// TIA Portal project "Demontagestation" (V17) (continued)
VERSION : 0.1
   VAR_INPUT
      Freigeben : Bool;   // "true", wenn der Funktionbaustein ausgeführt werden soll; bei "false werden die Ausgänge auf "Null" gesetzt
      Befehlsindex : USInt;   // Der Index zeigt auf einem Befehl, den der Greifer dann ausführen soll. {0 = FastStop, 1 = Stop, 2 = Quittierung, 3 = Referenzierung, 4 = Hubmessung, 5 = Greifen, 6 = Loslassen, 7 = Positionsfahrt, 8 = Relativfahrt}
      Kraftmodus : USInt;   // Der Wert (0 - 7) stellt die Art (Fast- oder Softgrip) und Kraft (100%, 75%, 50%, 25%) des Greifens ein (relevant bei Greifen).
      Außen_Innen : Bool;   // "true", wenn das Werkstück von innen gegriffen werden soll, sonst "false" (relevant bei Greifen und Loslassen)
      Zielposition : Real;   // Der Geifer positioniert sich nach dem vorgegebenen Positionswert (relevant bei Positions- und Relativfahrt).
   END_VAR
   VAR_OUTPUT
      Rückmeldung : String;   // Detaillierte Informationen über den Ausführungsstatus
      Fehler : Bool;   // "true", wenn im Prozess einen Fehler anliegt
      Fehlermeldung : String;   // Detaillierte Informationen über den Fehler.
      Hub_aktuell : Real;   // Der aktuelle Wert der Postition des Greifers
   END_VAR
   VAR_IN_OUT
      Ausführen : Bool;   // "true", um zu bestätigen, dass der Greifer aus den eingetragenen Daten den Befehl ausführen soll
   END_VAR
   VAR
      Befehlswert : Byte;   // Rohdatenwert eines Befehls
   END_VAR
   VAR_TEMP
      Prozessbit : Bool;   // "true", wenn der Befehl abgearbeitet ist
      Erfolg : Bool;   // "true", wenn der Befehl erfolgreich vollständig ausgeführt wurde
      Error : Bool;   // Quittierungspflichtige Fehler
      Spezifikationsfehler : Bool;   // Fehler, bei dem ein eingetragener Wert außerhalb des Gültigkeitsbereiches liegt
      Wartung : Bool;   // "true", wenn der Greifer gewartet werden muss
      Betrieb : Bool;   // "true", wenn der Greifer betriebsbereit ist
      Referenziert : Bool;   // "true", wenn der Greifer referenziert ist
   END_VAR
   VAR CONSTANT
      "BEGINN_E-ADRESSE" : Int := 39;   // Beginn der Eingangsadresse in Hardware-Konfiguration
      "BEGINN_A-ADRESSE" : Int := 29;   // Beginn der Eingangsadresse in Hardware-Konfiguration / Beginn der Ausgangsadresse in Hardware-Konfiguration
      NOTINDEX : USInt := 0;   // Index, der auf einem Notbefehl zuweist
      FEHLERWERT : Byte := -1;   // Wert, der statt auf einem Befehl einem Fehler weist.
      QUITTIERUNG : Byte := 16#1;   // Nach Beheben eines Fehlers wird der Greifer durch Quittieren des Fehlers vom Fehlerzustand in den normalen Betriebszustand versetzt.
      REFERENZIERUNG : Byte := 16#2;   // Beim Referenzieren wird die Nullposition festgelegt. Der Greifer fährt in eingestellter Referenzierrichtung bis zum mechanischen Endanschlag.
      HUBMESSUNG : Byte := 16#7;   // Bei der Hubmessung wird der maximale Hub des Greifers gegenüber der Referenzierposition festgelegt.
      GREIFEN : Byte := 16#4;   // Beim Greifen wird in Greifrichtung bis zum Anschlag gefahren und das Werkstück mit eingestellter Greifkraft gehalten.
      LOSLASSEN : Byte := 16#3;   // Beim Loslassen wird entgegen der Greifrichtung bis auf Endanschlag gefahren.
      POSITIONSFAHRT : Byte := 16#5;   // Der Geifer fährt auf die unter "Zielposition" angegebene Position.
      RELATIVFAHRT : Byte := 16#6;   // Der Geifer fährt auf eine Position, die von der letzten aktuellen Position mit einem relativen Abstand ermittelt wird.
      STOP : Byte := 16#8;   // Der Greifer wird geregelt in Stillstand versetzt.
      FASTSTOP : Byte := 16#0;   // Die elektrische Energieversorgung zum Aktor wird sofort unterbrochen, der Greifer wird ungesteuert stillgesetzt.
   END_VAR
BEGIN

REGION Network 1: Befehlszuweisung
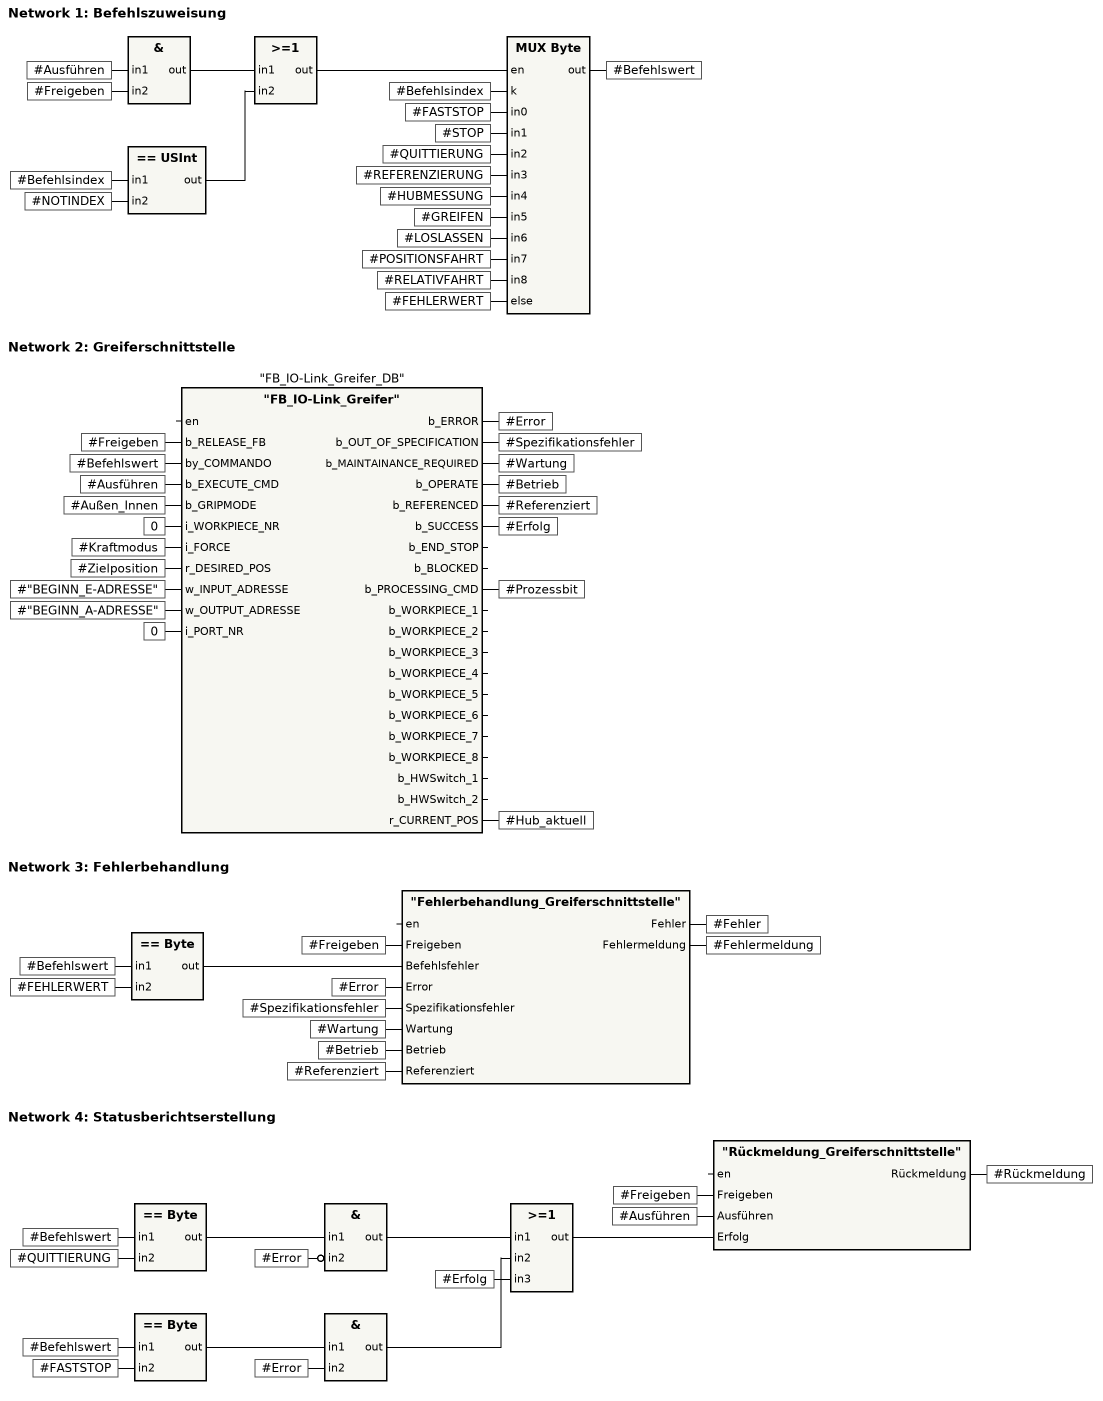
   // no SCL statement known for Mux: written as a call
   IF (#Ausführen AND #Freigeben) OR (#Befehlsindex = #NOTINDEX) THEN
       Mux(k := #Befehlsindex,
           in0 := #FASTSTOP,
           in1 := #STOP,
           in2 := #QUITTIERUNG,
           in3 := #REFERENZIERUNG,
           in4 := #HUBMESSUNG,
           in5 := #GREIFEN,
           in6 := #LOSLASSEN,
           in7 := #POSITIONSFAHRT,
           in8 := #RELATIVFAHRT,
           "else" := #FEHLERWERT,
           out => #Befehlswert);
   END_IF;
END_REGION

REGION Network 2: Greiferschnittstelle
   "FB_IO-Link_Greifer_DB"(b_RELEASE_FB := #Freigeben,   // "FB_IO-Link_Greifer"
                           by_COMMANDO := #Befehlswert,
                           b_EXECUTE_CMD := #Ausführen,
                           b_GRIPMODE := #Außen_Innen,
                           i_WORKPIECE_NR := 0,
                           i_FORCE := #Kraftmodus,
                           r_DESIRED_POS := #Zielposition,
                           w_INPUT_ADRESSE := #"BEGINN_E-ADRESSE",
                           w_OUTPUT_ADRESSE := #"BEGINN_A-ADRESSE",
                           i_PORT_NR := 0,
                           b_ERROR => #Error,
                           b_OUT_OF_SPECIFICATION => #Spezifikationsfehler,
                           b_MAINTAINANCE_REQUIRED => #Wartung,
                           b_OPERATE => #Betrieb,
                           b_REFERENCED => #Referenziert,
                           b_SUCCESS => #Erfolg,
                           b_PROCESSING_CMD => #Prozessbit,
                           r_CURRENT_POS => #Hub_aktuell);
END_REGION

REGION Network 3: Fehlerbehandlung
   "Fehlerbehandlung_Greiferschnittstelle"(Freigeben := #Freigeben,
                           Befehlsfehler := #Befehlswert = #FEHLERWERT,
                           Error := #Error,
                           Spezifikationsfehler := #Spezifikationsfehler,
                           Wartung := #Wartung,
                           Betrieb := #Betrieb,
                           Referenziert := #Referenziert,
                           Fehler => #Fehler,
                           Fehlermeldung => #Fehlermeldung);
END_REGION

REGION Network 4: Statusberichtserstellung
   "Rückmeldung_Greiferschnittstelle"(Freigeben := #Freigeben,
                           Ausführen := #Ausführen,
                           Erfolg := ((#Befehlswert = #QUITTIERUNG) AND NOT #Error) OR ((#Befehlswert = #FASTSTOP) AND #Error) OR #Erfolg,
                           Rückmeldung => #Rückmeldung);
END_REGION

REGION Network 5: Ausführungsende
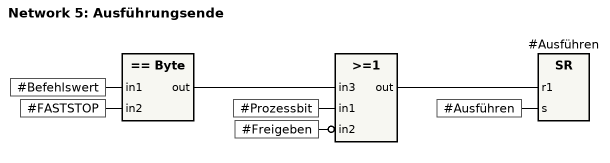
   IF #Ausführen THEN
       #Ausführen := TRUE;   // SR flip-flop
   END_IF;
   IF (#Befehlswert = #FASTSTOP) OR #Prozessbit OR NOT #Freigeben THEN #Ausführen := FALSE; END_IF;
END_REGION
END_FUNCTION_BLOCK

FUNCTION "Meldung_Sprachzuweisung" : Void   // FC1, FBD
{ S7_Optimized_Access := 'TRUE' }
VERSION : 0.1
   VAR_INPUT
      Meldung_Deutsch : String;   // Meldung auf Deutsch
      Meldung_Englisch : String;   // Meldung auf Englisch
   END_VAR
   VAR_OUTPUT
      Meldung : String;   // Meldung in der eingestellten Sprache
   END_VAR
   VAR CONSTANT
      SPRACHINDEX : UInt := 1;   // 0 = Deutsch, 1 = Englisch
      INDEX_DEUTSCH : UInt := 0;   // Indexwert für Deutsch
      INDEX_ENGLISCH : UInt := 1;   // Indexwert für Englisch
   END_VAR
BEGIN

REGION Network 1: Zuweisung der deutschen Meldung
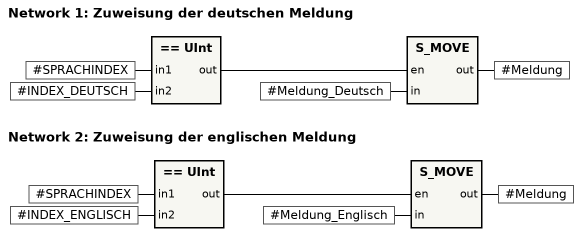
   IF #SPRACHINDEX = #INDEX_DEUTSCH THEN #Meldung := #Meldung_Deutsch; END_IF;
END_REGION

REGION Network 2: Zuweisung der englischen Meldung
   IF #SPRACHINDEX = #INDEX_ENGLISCH THEN #Meldung := #Meldung_Englisch; END_IF;
END_REGION
END_FUNCTION

FUNCTION "Fehlerbehandlung_Greiferschnittstelle" : Void   // FC6, FBD
{ S7_Optimized_Access := 'TRUE' }
VERSION : 0.1
   VAR_INPUT
      Freigeben : Bool;   // "true", wenn der Funktionbaustein ausgeführt werden soll; bei "false werden die Ausgänge auf "Null" gesetzt
      Befehlsfehler : Bool;   // Fehler, bei dem der eingetragene Befehlsindex keinen Befehl zugeordnet werden kann
      Error : Bool;   // Quittierungspflichtige Fehler
      Spezifikationsfehler : Bool;   // Fehler, bei dem ein eingetragener Wert außerhalb des Gültigkeitsbereiches liegt
      Wartung : Bool;   // "true", wenn der Greifer gewartet werden muss
      Betrieb : Bool;   // "true", wenn der Greifer betriebsbereit ist
      Referenziert : Bool;   // "true", wenn der Greifer referenziert ist
   END_VAR
   VAR_OUTPUT
      Fehler : Bool;   // "true", wenn im Prozess einen Fehler anliegt
      Fehlermeldung : String;   // Detaillierte Darstellung des Fehlers (nur relevant bei einem Fehler)
   END_VAR
   VAR_TEMP
      Falscher_Befehlsindex : String;   // Platzhalter für die Zuweisung der entsprechenden Meldung in der eingestellten Sprache
      Fehler_quittieren : String;   // Platzhalter für die Zuweisung der entsprechenden Meldung in der eingestellten Sprache
      Wert_ungültig : String;   // Platzhalter für die Zuweisung der entsprechenden Meldung in der eingestellten Sprache
      Wartung_nötig : String;   // Platzhalter für die Zuweisung der entsprechenden Meldung in der eingestellten Sprache
      Nicht_betriebsbereit : String;   // Platzhalter für die Zuweisung der entsprechenden Meldung in der eingestellten Sprache
      Nicht_referenziert : String;   // Platzhalter für die Zuweisung der entsprechenden Meldung in der eingestellten Sprache
   END_VAR
   VAR CONSTANT
      KEINE_MELDUNG : String := '';   // Leerer Text, um die vorherige Meldung zu löschen
      FALSCHER_BEFEHLSINDEX_D : String := 'Befehlsindex_nur_0-8_gueltig!';   // Fehlermeldung bei einer falschen Eingabe des Befehlsindexes (Deutsch)
      FALSCHER_BEFEHLSINDEX_E : String := 'Command_Index_only_0-8_valid!';   // Fehlermeldung bei einer falschen Eingabe des Befehlsindexes (Englisch)
      FEHLER_QUITTIEREN_D : String := 'Fehler_mit_"Quittierung"_aufheben!';   // Fehlermeldung bei einem Fehler, der zu quittieren ist (Deutsch)
      FEHLER_QUITTIEREN_E : String := 'Error_canceling_with_"Acknowledge"!';   // Fehlermeldung bei einem Fehler, der zu quittieren ist (Englisch)
      WERT_UNGÜLTIG_D : String := 'Ein_Wert_nicht_gueltig!';   // Fehlermeldung bei einem eingetragenen Wert, der außerhalb seines Gültigkeitsbereiches liegt (Deutsch)
      WERT_UNGÜLTIG_E : String := 'A_value_not_valid!';   // Fehlermeldung bei einem eingetragenen Wert, der außerhalb seines Gültigkeitsbereiches liegt (Englisch)
      WARTUNG_NÖTIG_D : String := 'Greifer_muss_gewartet_werden!';   // Fehlermeldung, wenn der Greifer gewartet werden muss (Deutsch)
      WARTUNG_NÖTIG_E : String := 'Gripper_requires_maintenance!';   // Fehlermeldung, wenn der Greifer gewartet werden muss (Englisch)
      NICHT_BETRIEBSBEREIT_D : String := 'Greifer_nicht_betriebsbereit!';   // Fehlermeldung, wenn der Greifer noch nicht betriebsbereit ist (Deutsch)
      NICHT_BETRIEBSBEREIT_E : String := 'Gripper_not_ready!';   // Fehlermeldung, wenn der Greifer noch nicht betriebsbereit ist (Englisch)
      NICHT_REFERENZIERT_D : String := 'Greifer_muss_referenziert_werden!';   // Fehlermeldung, wenn der Greifer noch nicht referenziert ist (Deutsch)
      NICHT_REFERENZIERT_E : String := 'Gripper_must_be_referenced!';   // Fehlermeldung, wenn der Greifer noch nicht referenziert ist (Englisch)
   END_VAR
   VAR_TEMP   // added for the SCL form of the ladder/FBD networks
      _w1 : Bool;
   END_VAR
BEGIN

REGION Network 1: Fehlersignal
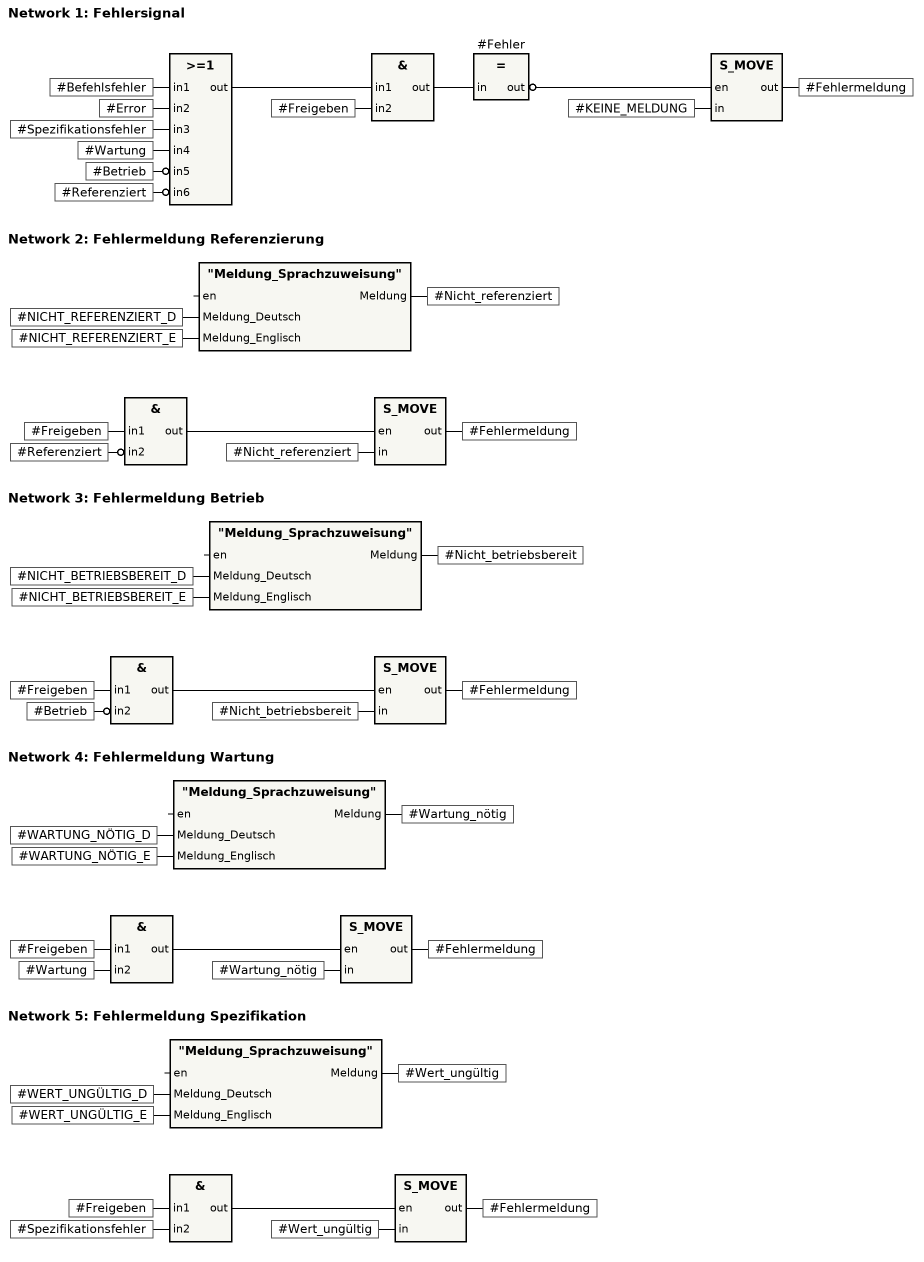
   #_w1 := (#Befehlsfehler OR #Error OR #Spezifikationsfehler OR #Wartung OR NOT #Betrieb OR NOT #Referenziert) AND #Freigeben;
   #Fehler := #_w1;
   IF NOT #_w1 THEN #Fehlermeldung := #KEINE_MELDUNG; END_IF;
END_REGION

REGION Network 2: Fehlermeldung Referenzierung
   "Meldung_Sprachzuweisung"(Meldung_Deutsch := #NICHT_REFERENZIERT_D,
                           Meldung_Englisch := #NICHT_REFERENZIERT_E,
                           Meldung => #Nicht_referenziert);
   IF #Freigeben AND NOT #Referenziert THEN #Fehlermeldung := #Nicht_referenziert; END_IF;
END_REGION

REGION Network 3: Fehlermeldung Betrieb
   "Meldung_Sprachzuweisung"(Meldung_Deutsch := #NICHT_BETRIEBSBEREIT_D,
                           Meldung_Englisch := #NICHT_BETRIEBSBEREIT_E,
                           Meldung => #Nicht_betriebsbereit);
   IF #Freigeben AND NOT #Betrieb THEN #Fehlermeldung := #Nicht_betriebsbereit; END_IF;
END_REGION

REGION Network 4: Fehlermeldung Wartung
   "Meldung_Sprachzuweisung"(Meldung_Deutsch := #WARTUNG_NÖTIG_D,
                           Meldung_Englisch := #WARTUNG_NÖTIG_E,
                           Meldung => #Wartung_nötig);
   IF #Freigeben AND #Wartung THEN #Fehlermeldung := #Wartung_nötig; END_IF;
END_REGION

REGION Network 5: Fehlermeldung Spezifikation
   "Meldung_Sprachzuweisung"(Meldung_Deutsch := #WERT_UNGÜLTIG_D,
                           Meldung_Englisch := #WERT_UNGÜLTIG_E,
                           Meldung => #Wert_ungültig);
   IF #Freigeben AND #Spezifikationsfehler THEN #Fehlermeldung := #Wert_ungültig; END_IF;
END_REGION

REGION Network 6: Fehlermeldung Error
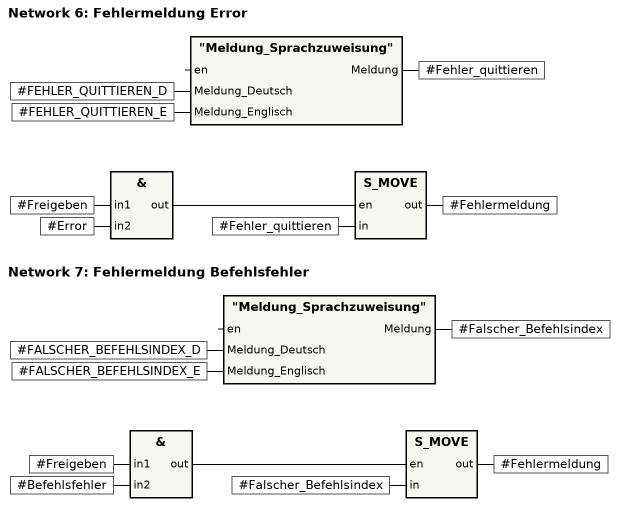
   "Meldung_Sprachzuweisung"(Meldung_Deutsch := #FEHLER_QUITTIEREN_D,
                           Meldung_Englisch := #FEHLER_QUITTIEREN_E,
                           Meldung => #Fehler_quittieren);
   IF #Freigeben AND #Error THEN #Fehlermeldung := #Fehler_quittieren; END_IF;
END_REGION

REGION Network 7: Fehlermeldung Befehlsfehler
   "Meldung_Sprachzuweisung"(Meldung_Deutsch := #FALSCHER_BEFEHLSINDEX_D,
                           Meldung_Englisch := #FALSCHER_BEFEHLSINDEX_E,
                           Meldung => #Falscher_Befehlsindex);
   IF #Freigeben AND #Befehlsfehler THEN #Fehlermeldung := #Falscher_Befehlsindex; END_IF;
END_REGION
END_FUNCTION

FUNCTION "Rückmeldung_Greiferschnittstelle" : Void   // FC7, FBD
{ S7_Optimized_Access := 'TRUE' }
VERSION : 0.1
   VAR_INPUT
      Freigeben : Bool;   // "true", wenn der Funktionbaustein ausgeführt werden soll; bei "false werden die Ausgänge auf "Null" gesetzt
      Ausführen : Bool;   // "true", um zu bestätigen, dass der Greifer aus den eingetragenen Daten den Befehl ausführen soll
      Erfolg : Bool;   // "true", wenn der Befehl erfolgreich vollständig ausgeführt wurde
   END_VAR
   VAR_OUTPUT
      Rückmeldung : String;   // Detaillierte Informationen über den Ausführungsstatus
   END_VAR
   VAR_TEMP
      In_Prozess : String;   // Platzhalter für die Zuweisung der entsprechenden Meldung in der eingestellten Sprache
      Erfolgreich : String;   // Platzhalter für die Zuweisung der entsprechenden Meldung in der eingestellten Sprache
      Nicht_erfolgreich : String;   // Platzhalter für die Zuweisung der entsprechenden Meldung in der eingestellten Sprache
   END_VAR
   VAR CONSTANT
      KEINE_MELDUNG : String := '';   // Leerer Text, um die vorherige Meldung zu löschen
      IN_PROZESS_D : String := 'Befehl_in_Arbeit!';   // Rückmeldung, wenn der Befehl gerade abgearbeitet wird (Deutsch)
      IN_PROZESS_E : String := 'Command_in_progress!';   // Rückmeldung, wenn der Befehl gerade abgearbeitet wird (Englisch)
      ERFOLGREICH_D : String := 'Befehl_ausgefuehrt!';   // Rückmeldung, wenn der Befehl vollständig ausgeführt wurde (Deutsch)
      ERFOLGREICH_E : String := 'Command_executed!';   // Rückmeldung, wenn der Befehl vollständig ausgeführt wurde (Englisch)
      NICHT_ERFOLGREICH_D : String := 'Befehl_nicht_ausgefuehrt!';   // Rückmeldung, wenn der Befhel nicht vollständig ausgeführt wurde (Deutsch)
      NICHT_ERFOLGREICH_E : String := 'Command_not_executed!';   // Rückmeldung, wenn der Befhel nicht vollständig ausgeführt wurde (Englisch)
   END_VAR
   VAR_TEMP   // added for the SCL form of the ladder/FBD networks
      _w1 : Bool;
   END_VAR
BEGIN

REGION Network 1: Meldung leeren
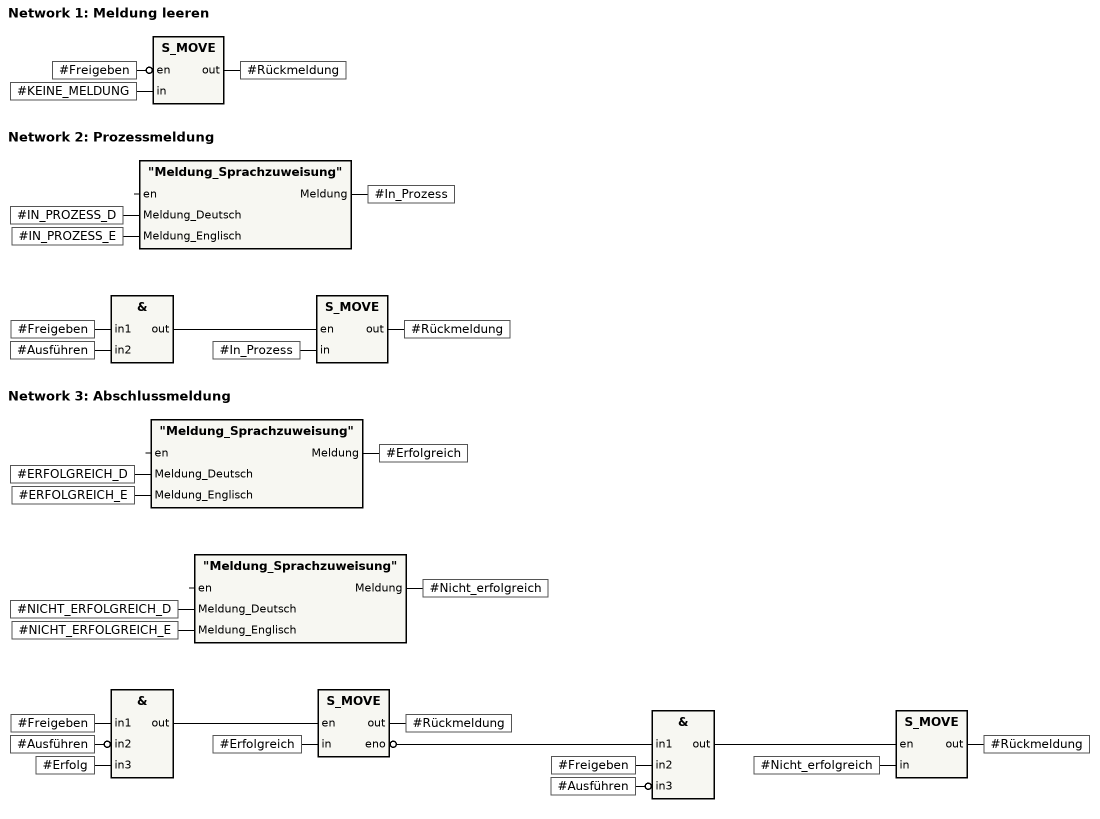
   IF NOT #Freigeben THEN #Rückmeldung := #KEINE_MELDUNG; END_IF;
END_REGION

REGION Network 2: Prozessmeldung
   "Meldung_Sprachzuweisung"(Meldung_Deutsch := #IN_PROZESS_D,
                           Meldung_Englisch := #IN_PROZESS_E,
                           Meldung => #In_Prozess);
   IF #Freigeben AND #Ausführen THEN #Rückmeldung := #In_Prozess; END_IF;
END_REGION

REGION Network 3: Abschlussmeldung
   "Meldung_Sprachzuweisung"(Meldung_Deutsch := #ERFOLGREICH_D,
                           Meldung_Englisch := #ERFOLGREICH_E,
                           Meldung => #Erfolgreich);
   "Meldung_Sprachzuweisung"(Meldung_Deutsch := #NICHT_ERFOLGREICH_D,
                           Meldung_Englisch := #NICHT_ERFOLGREICH_E,
                           Meldung => #Nicht_erfolgreich);
   #_w1 := #Freigeben AND NOT #Ausführen AND #Erfolg;
   IF #_w1 THEN #Rückmeldung := #Erfolgreich; END_IF;
   IF NOT #_w1 AND #Freigeben AND NOT #Ausführen THEN #Rückmeldung := #Nicht_erfolgreich; END_IF;
END_REGION
END_FUNCTION

// folder: Pneumatik

FUNCTION_BLOCK "Luftdrucksteuerung"   // FB5, FBD
{ S7_Optimized_Access := 'TRUE' }
VERSION : 0.1
   VAR_INPUT
      "Hand/Automatik" : Bool;
      "Ist-Luftdruck" : Int;
      "Soll-Luftdruck" : Real;
      "Luftdruck erhöhen" : Bool;
      "Luftdruck senken" : Bool;
   END_VAR
   VAR_OUTPUT
      Ausgabeluftdruck : Int;
   END_VAR
   VAR
      Handbetrieb : Bool;
      Automatikbetrieb : Bool;
      "Flanke Luftdruck erhöhen" : Bool;
      "Flanke Luftdruck Senken" : Bool;
      "Ist-Luftdruck Skaliert" : Int;
      "Ist-Luftdruck Normiert" : Real;
      "Ausgabeluftdruck unskaliert" : Int;
      "Ausgabedruck unnomiert" : Real;
      "Soll-Luftdruck Int" : Int;
   END_VAR
   VAR_TEMP   // added for the SCL form of the ladder/FBD networks
      _w1 : Bool;
   END_VAR
BEGIN

REGION Network 1: Betriebsart
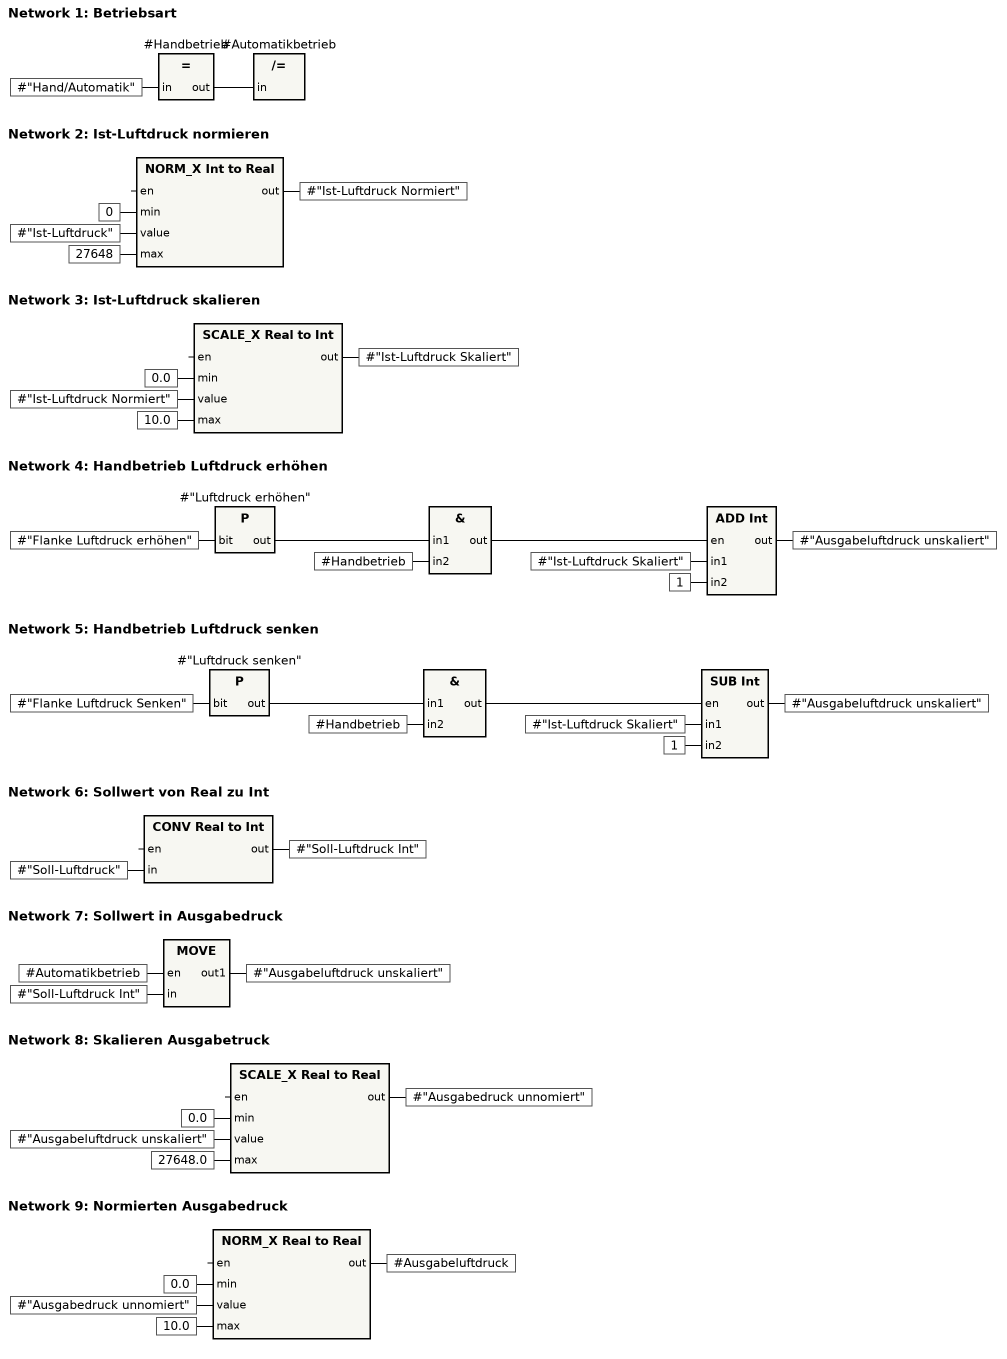
   #Handbetrieb := #"Hand/Automatik";
   #Automatikbetrieb := NOT #"Hand/Automatik";
END_REGION

REGION Network 2: Ist-Luftdruck normieren
   #"Ist-Luftdruck Normiert" := NORM_X(MIN := 0, VALUE := #"Ist-Luftdruck", MAX := 27648);
END_REGION

REGION Network 3: Ist-Luftdruck skalieren
   #"Ist-Luftdruck Skaliert" := SCALE_X(MIN := 0.0, VALUE := #"Ist-Luftdruck Normiert", MAX := 10.0);
END_REGION

REGION Network 4: Handbetrieb Luftdruck erhöhen
   #_w1 := #"Luftdruck erhöhen" AND NOT #"Flanke Luftdruck erhöhen";   // rising edge of #"Luftdruck erhöhen"
   #"Flanke Luftdruck erhöhen" := #"Luftdruck erhöhen";
   IF #_w1 AND #Handbetrieb THEN #"Ausgabeluftdruck unskaliert" := #"Ist-Luftdruck Skaliert" + 1; END_IF;
END_REGION

REGION Network 5: Handbetrieb Luftdruck senken
   #_w1 := #"Luftdruck senken" AND NOT #"Flanke Luftdruck Senken";   // rising edge of #"Luftdruck senken"
   #"Flanke Luftdruck Senken" := #"Luftdruck senken";
   IF #_w1 AND #Handbetrieb THEN #"Ausgabeluftdruck unskaliert" := #"Ist-Luftdruck Skaliert" - 1; END_IF;
END_REGION

REGION Network 6: Sollwert von Real zu Int
   #"Soll-Luftdruck Int" := REAL_TO_INT(#"Soll-Luftdruck");
END_REGION

REGION Network 7: Sollwert in Ausgabedruck
   IF #Automatikbetrieb THEN #"Ausgabeluftdruck unskaliert" := #"Soll-Luftdruck Int"; END_IF;
END_REGION

REGION Network 8: Skalieren Ausgabetruck
   #"Ausgabedruck unnomiert" := SCALE_X(MIN := 0.0, VALUE := #"Ausgabeluftdruck unskaliert", MAX := 27648.0);
END_REGION

REGION Network 9: Normierten Ausgabedruck
   #Ausgabeluftdruck := NORM_X(MIN := 0.0, VALUE := #"Ausgabedruck unnomiert", MAX := 10.0);
END_REGION
END_FUNCTION_BLOCK